// TIA Portal project "Hydroelectric Power Plant" (V20) (continued)
VERSION : 0.1
   VAR
      Os1 : Bool;
      Os2 : Bool;
      Os3 : Bool;
      Os4 : Bool;
      Os5 : Bool;
      Os6 : Bool;
      Os7 : Bool;
      Os8 : Bool;
      Os9 : Bool;
      Os10 : Bool;
      Os11 : Bool;
      Os12 : Bool;
   END_VAR
   VAR_TEMP   // added for the SCL form of the ladder/FBD networks
      _w1 : Bool;
      _w2 : Bool;
      _w3 : Bool;
   END_VAR
BEGIN

REGION Network 1
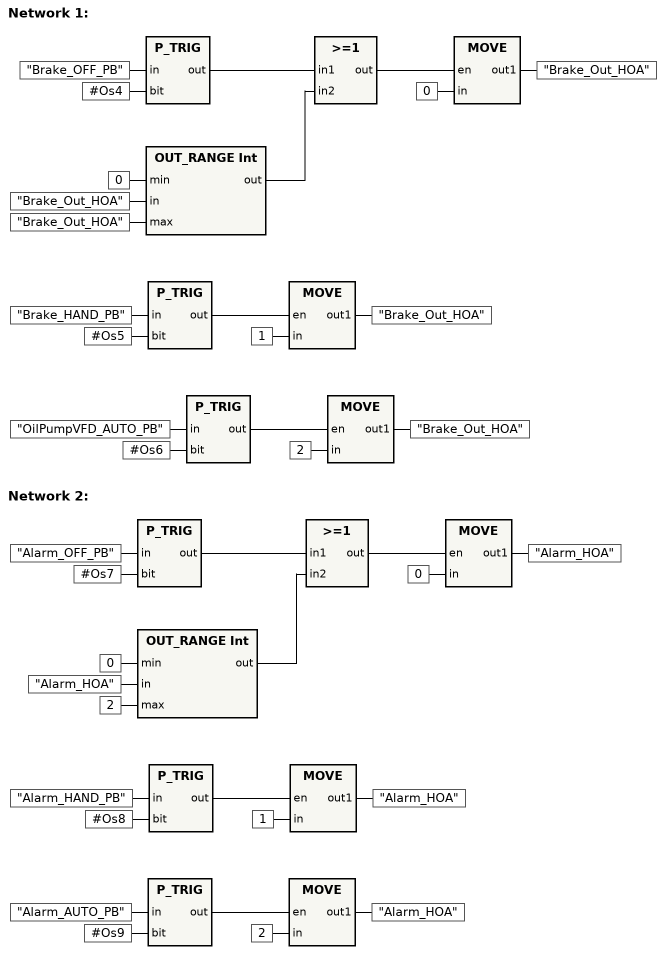
   #_w1 := "Brake_OFF_PB" AND NOT #Os4;   // rising edge
   #Os4 := "Brake_OFF_PB";
   IF #_w1 OR ("Brake_Out_HOA" < 0) OR ("Brake_Out_HOA" > "Brake_Out_HOA") THEN "Brake_Out_HOA" := 0; END_IF;
   #_w2 := "Brake_HAND_PB" AND NOT #Os5;   // rising edge
   #Os5 := "Brake_HAND_PB";
   IF #_w2 THEN "Brake_Out_HOA" := 1; END_IF;
   #_w3 := "OilPumpVFD_AUTO_PB" AND NOT #Os6;   // rising edge
   #Os6 := "OilPumpVFD_AUTO_PB";
   IF #_w3 THEN "Brake_Out_HOA" := 2; END_IF;
END_REGION

REGION Network 2
   #_w1 := "Alarm_OFF_PB" AND NOT #Os7;   // rising edge
   #Os7 := "Alarm_OFF_PB";
   IF #_w1 OR ("Alarm_HOA" < 0) OR ("Alarm_HOA" > 2) THEN "Alarm_HOA" := 0; END_IF;
   #_w2 := "Alarm_HAND_PB" AND NOT #Os8;   // rising edge
   #Os8 := "Alarm_HAND_PB";
   IF #_w2 THEN "Alarm_HOA" := 1; END_IF;
   #_w3 := "Alarm_AUTO_PB" AND NOT #Os9;   // rising edge
   #Os9 := "Alarm_AUTO_PB";
   IF #_w3 THEN "Alarm_HOA" := 2; END_IF;
END_REGION

REGION Network 3
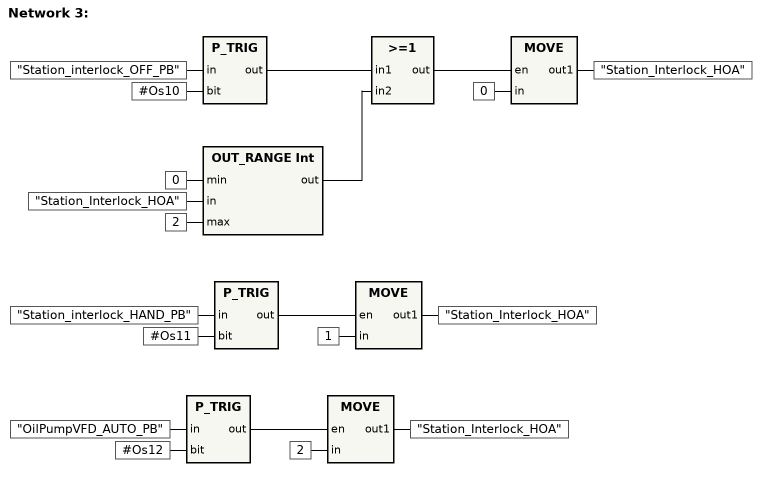
   #_w1 := "Station_interlock_OFF_PB" AND NOT #Os10;   // rising edge
   #Os10 := "Station_interlock_OFF_PB";
   IF #_w1 OR ("Station_Interlock_HOA" < 0) OR ("Station_Interlock_HOA" > 2) THEN
       "Station_Interlock_HOA" := 0;
   END_IF;
   #_w2 := "Station_interlock_HAND_PB" AND NOT #Os11;   // rising edge
   #Os11 := "Station_interlock_HAND_PB";
   IF #_w2 THEN "Station_Interlock_HOA" := 1; END_IF;
   #_w3 := "OilPumpVFD_AUTO_PB" AND NOT #Os12;   // rising edge
   #Os12 := "OilPumpVFD_AUTO_PB";
   IF #_w3 THEN "Station_Interlock_HOA" := 2; END_IF;
END_REGION
END_FUNCTION_BLOCK

FUNCTION_BLOCK "Alarm_FBD"   // FB11, FBD
{ S7_Optimized_Access := 'TRUE' }
VERSION : 0.1
   VAR
      OS1 : Bool;
      OS2 : Bool;
      OS3 : Bool;
      OS4 : Bool;
      OS5 : Bool;
      OS6 : Bool;
      OS7 : Bool;
      on8 : Bool;
   END_VAR
   VAR_TEMP
      tp1 : Int;
      OLFD : Time;
      tp2 : Int;
      OCD : Time;
      tp3 : Int;
      tp4 : Int;
      tp5 : Int;
      tp6 : Int;
      tp7 : Int;
      HOT : Time;
      OHF : Time;
      ROS : Time;
      BF : Time;
      AlarmTrigger : Bool;
   END_VAR
   VAR_TEMP   // added for the SCL form of the ladder/FBD networks
      _w1 : Bool;
   END_VAR
BEGIN

REGION Network 1: Oil_Low_Flow_Alarm
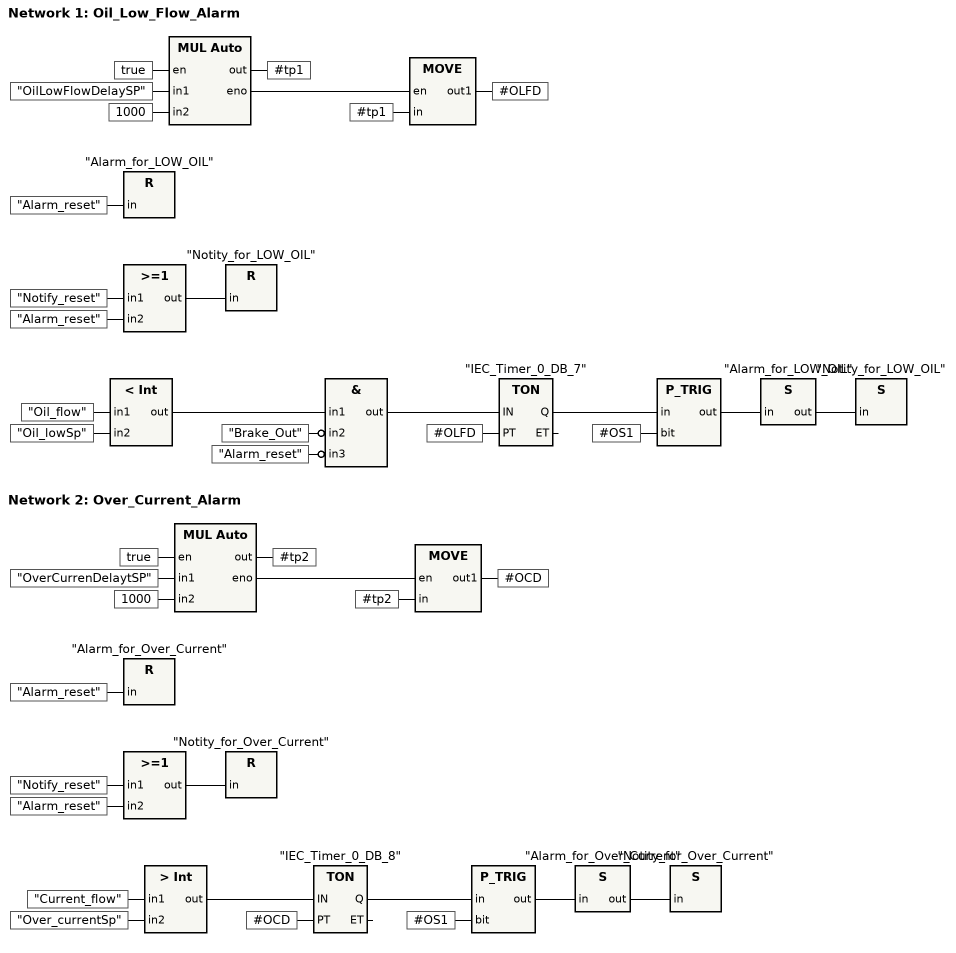
   IF true THEN
       #tp1 := "OilLowFlowDelaySP" * 1000;
       #OLFD := #tp1;
   END_IF;
   IF "Alarm_reset" THEN "Alarm_for_LOW_OIL" := FALSE; END_IF;
   IF "Notify_reset" OR "Alarm_reset" THEN "Notity_for_LOW_OIL" := FALSE; END_IF;
   "IEC_Timer_0_DB_7".TON(IN := ("Oil_flow" < "Oil_lowSp") AND NOT "Brake_Out" AND NOT "Alarm_reset",
                          PT := #OLFD);
   #_w1 := "IEC_Timer_0_DB_7".Q AND NOT #OS1;   // rising edge
   #OS1 := "IEC_Timer_0_DB_7".Q;
   IF #_w1 THEN
       "Alarm_for_LOW_OIL" := TRUE;
       "Notity_for_LOW_OIL" := TRUE;
   END_IF;
END_REGION

REGION Network 2: Over_Current_Alarm
   IF true THEN
       #tp2 := "OverCurrenDelaytSP" * 1000;
       #OCD := #tp2;
   END_IF;
   IF "Alarm_reset" THEN "Alarm_for_Over_Current" := FALSE; END_IF;
   IF "Notify_reset" OR "Alarm_reset" THEN "Notity_for_Over_Current" := FALSE; END_IF;
   "IEC_Timer_0_DB_8".TON(IN := "Current_flow" > "Over_currentSp", PT := #OCD);
   #_w1 := "IEC_Timer_0_DB_8".Q AND NOT #OS1;   // rising edge
   #OS1 := "IEC_Timer_0_DB_8".Q;
   IF #_w1 THEN
       "Alarm_for_Over_Current" := TRUE;
       "Notity_for_Over_Current" := TRUE;
   END_IF;
END_REGION

REGION Network 3: High_Oil_Temp_Alarm
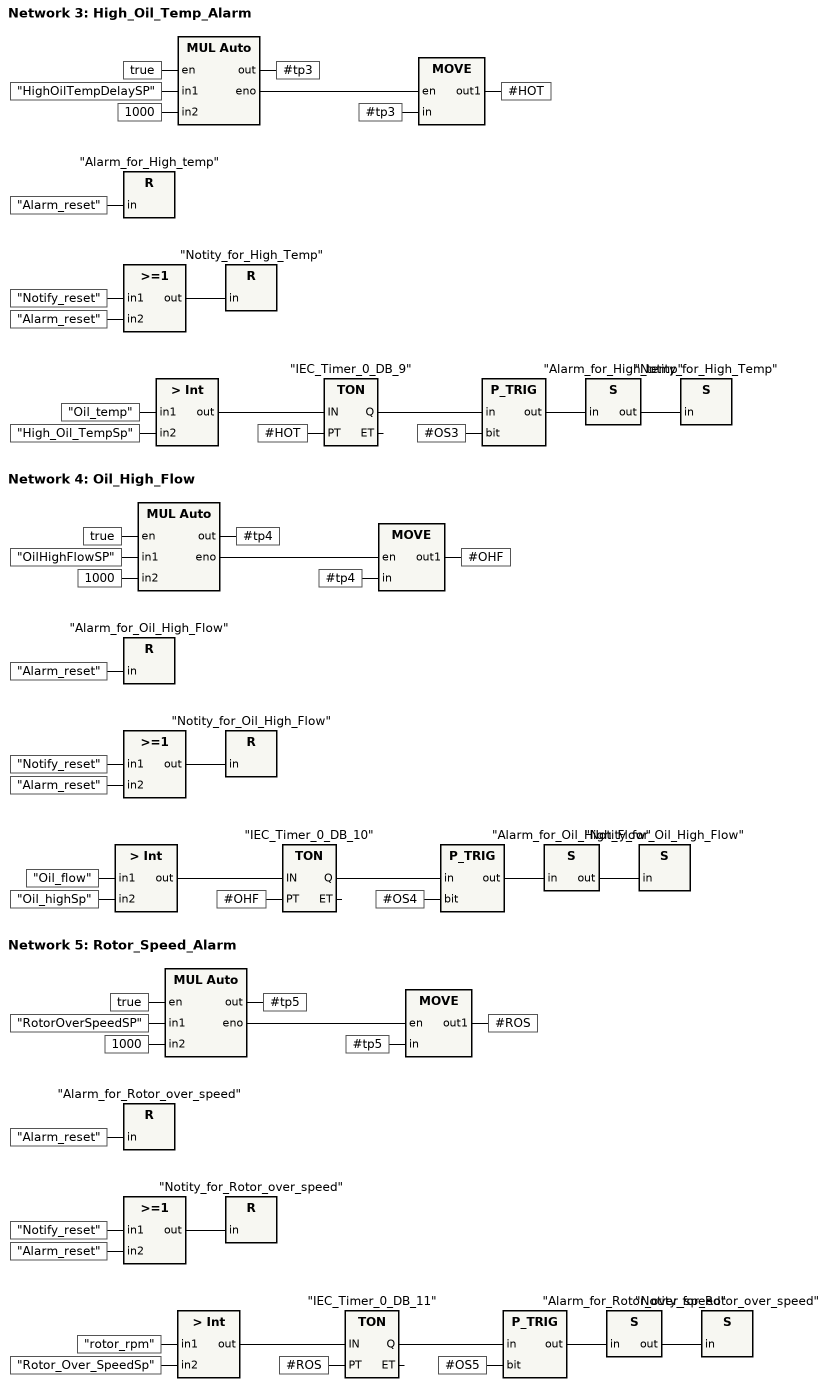
   IF true THEN
       #tp3 := "HighOilTempDelaySP" * 1000;
       #HOT := #tp3;
   END_IF;
   IF "Alarm_reset" THEN "Alarm_for_High_temp" := FALSE; END_IF;
   IF "Notify_reset" OR "Alarm_reset" THEN "Notity_for_High_Temp" := FALSE; END_IF;
   "IEC_Timer_0_DB_9".TON(IN := "Oil_temp" > "High_Oil_TempSp", PT := #HOT);
   #_w1 := "IEC_Timer_0_DB_9".Q AND NOT #OS3;   // rising edge
   #OS3 := "IEC_Timer_0_DB_9".Q;
   IF #_w1 THEN
       "Alarm_for_High_temp" := TRUE;
       "Notity_for_High_Temp" := TRUE;
   END_IF;
END_REGION

REGION Network 4: Oil_High_Flow
   IF true THEN
       #tp4 := "OilHighFlowSP" * 1000;
       #OHF := #tp4;
   END_IF;
   IF "Alarm_reset" THEN "Alarm_for_Oil_High_Flow" := FALSE; END_IF;
   IF "Notify_reset" OR "Alarm_reset" THEN "Notity_for_Oil_High_Flow" := FALSE; END_IF;
   "IEC_Timer_0_DB_10".TON(IN := "Oil_flow" > "Oil_highSp", PT := #OHF);
   #_w1 := "IEC_Timer_0_DB_10".Q AND NOT #OS4;   // rising edge
   #OS4 := "IEC_Timer_0_DB_10".Q;
   IF #_w1 THEN
       "Alarm_for_Oil_High_Flow" := TRUE;
       "Notity_for_Oil_High_Flow" := TRUE;
   END_IF;
END_REGION

REGION Network 5: Rotor_Speed_Alarm
   IF true THEN
       #tp5 := "RotorOverSpeedSP" * 1000;
       #ROS := #tp5;
   END_IF;
   IF "Alarm_reset" THEN "Alarm_for_Rotor_over_speed" := FALSE; END_IF;
   IF "Notify_reset" OR "Alarm_reset" THEN "Notity_for_Rotor_over_speed" := FALSE; END_IF;
   "IEC_Timer_0_DB_11".TON(IN := "rotor_rpm" > "Rotor_Over_SpeedSp", PT := #ROS);
   #_w1 := "IEC_Timer_0_DB_11".Q AND NOT #OS5;   // rising edge
   #OS5 := "IEC_Timer_0_DB_11".Q;
   IF #_w1 THEN
       "Alarm_for_Rotor_over_speed" := TRUE;
       "Notity_for_Rotor_over_speed" := TRUE;
   END_IF;
END_REGION

REGION Network 6: Brake_Failure_Alarm
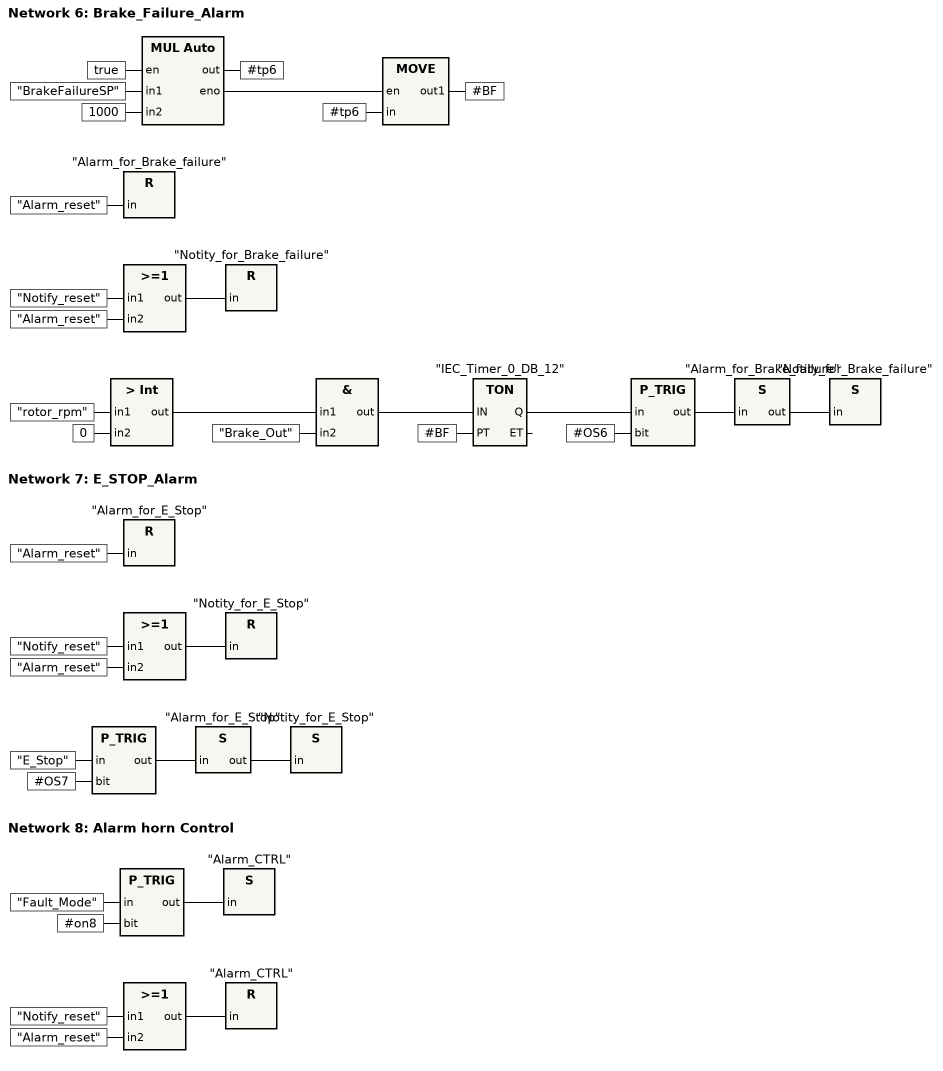
   IF true THEN
       #tp6 := "BrakeFailureSP" * 1000;
       #BF := #tp6;
   END_IF;
   IF "Alarm_reset" THEN "Alarm_for_Brake_failure" := FALSE; END_IF;
   IF "Notify_reset" OR "Alarm_reset" THEN "Notity_for_Brake_failure" := FALSE; END_IF;
   "IEC_Timer_0_DB_12".TON(IN := ("rotor_rpm" > 0) AND "Brake_Out", PT := #BF);
   #_w1 := "IEC_Timer_0_DB_12".Q AND NOT #OS6;   // rising edge
   #OS6 := "IEC_Timer_0_DB_12".Q;
   IF #_w1 THEN
       "Alarm_for_Brake_failure" := TRUE;
       "Notity_for_Brake_failure" := TRUE;
   END_IF;
END_REGION

REGION Network 7: E_STOP_Alarm
   IF "Alarm_reset" THEN "Alarm_for_E_Stop" := FALSE; END_IF;
   IF "Notify_reset" OR "Alarm_reset" THEN "Notity_for_E_Stop" := FALSE; END_IF;
   #_w1 := "E_Stop" AND NOT #OS7;   // rising edge
   #OS7 := "E_Stop";
   IF #_w1 THEN
       "Alarm_for_E_Stop" := TRUE;
       "Notity_for_E_Stop" := TRUE;
   END_IF;
END_REGION

REGION Network 8: Alarm horn Control
   #_w1 := "Fault_Mode" AND NOT #on8;   // rising edge
   #on8 := "Fault_Mode";
   IF #_w1 THEN "Alarm_CTRL" := TRUE; END_IF;
   IF "Notify_reset" OR "Alarm_reset" THEN "Alarm_CTRL" := FALSE; END_IF;
END_REGION
END_FUNCTION_BLOCK

FUNCTION_BLOCK "Modes_FBD"   // FB15, FBD
{ S7_Optimized_Access := 'TRUE' }
VERSION : 0.1
   VAR
      os1 : Bool;
      os2 : Bool;
      os3 : Bool;
      os4 : Bool;
      os5 : Bool;
      os6 : Bool;
   END_VAR
   VAR_TEMP
      ti1 : Time;
      tv2 : Int;
      tv1 : Int;
      ti2 : Time;
      ti3 : Time;
   END_VAR
   VAR_TEMP   // added for the SCL form of the ladder/FBD networks
      _w1 : Bool;
      _w2 : Bool;
      _w3 : Bool;
   END_VAR
BEGIN

REGION Network 1: WarmUp_Mode
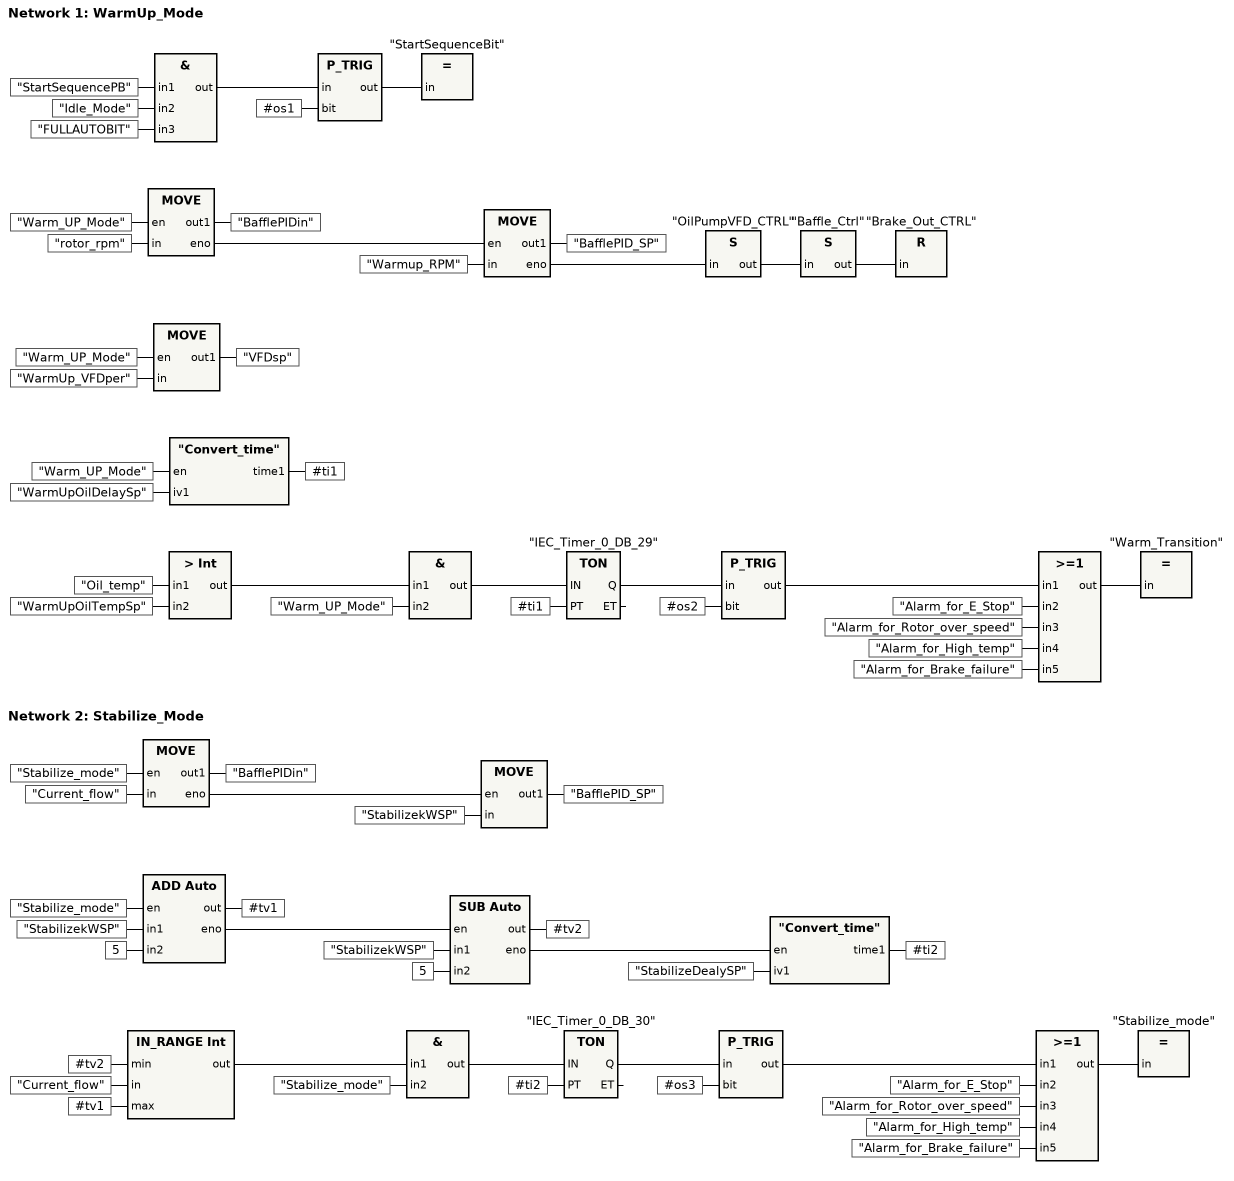
   #_w1 := "StartSequencePB" AND "Idle_Mode" AND "FULLAUTOBIT";
   #_w2 := #_w1 AND NOT #os1;   // rising edge
   #os1 := #_w1;
   "StartSequenceBit" := #_w2;
   IF "Warm_UP_Mode" THEN
       "BafflePIDin" := "rotor_rpm";
       "BafflePID_SP" := "Warmup_RPM";
       "OilPumpVFD_CTRL" := TRUE;
       "Baffle_Ctrl" := TRUE;
       "Brake_Out_CTRL" := FALSE;
       "VFDsp" := "WarmUp_VFDper";
       "Convert_time"(iv1 := "WarmUpOilDelaySp", time1 => #ti1);
   END_IF;
   "IEC_Timer_0_DB_29".TON(IN := ("Oil_temp" > "WarmUpOilTempSp") AND "Warm_UP_Mode", PT := #ti1);
   #_w3 := "IEC_Timer_0_DB_29".Q AND NOT #os2;   // rising edge
   #os2 := "IEC_Timer_0_DB_29".Q;
   "Warm_Transition" := #_w3 OR "Alarm_for_E_Stop" OR "Alarm_for_Rotor_over_speed" OR "Alarm_for_High_temp" OR "Alarm_for_Brake_failure";
END_REGION

REGION Network 2: Stabilize_Mode
   IF "Stabilize_mode" THEN
       "BafflePIDin" := "Current_flow";
       "BafflePID_SP" := "StabilizekWSP";
       #tv1 := "StabilizekWSP" + 5;
       #tv2 := "StabilizekWSP" - 5;
       "Convert_time"(iv1 := "StabilizeDealySP", time1 => #ti2);
   END_IF;
   "IEC_Timer_0_DB_30".TON(IN := (#tv2 <= "Current_flow") AND ("Current_flow" <= #tv1) AND "Stabilize_mode",
                           PT := #ti2);
   #_w1 := "IEC_Timer_0_DB_30".Q AND NOT #os3;   // rising edge
   #os3 := "IEC_Timer_0_DB_30".Q;
   "Stabilize_mode" := #_w1 OR "Alarm_for_E_Stop" OR "Alarm_for_Rotor_over_speed" OR "Alarm_for_High_temp" OR "Alarm_for_Brake_failure";
END_REGION

REGION Network 3: Gereration_Mode
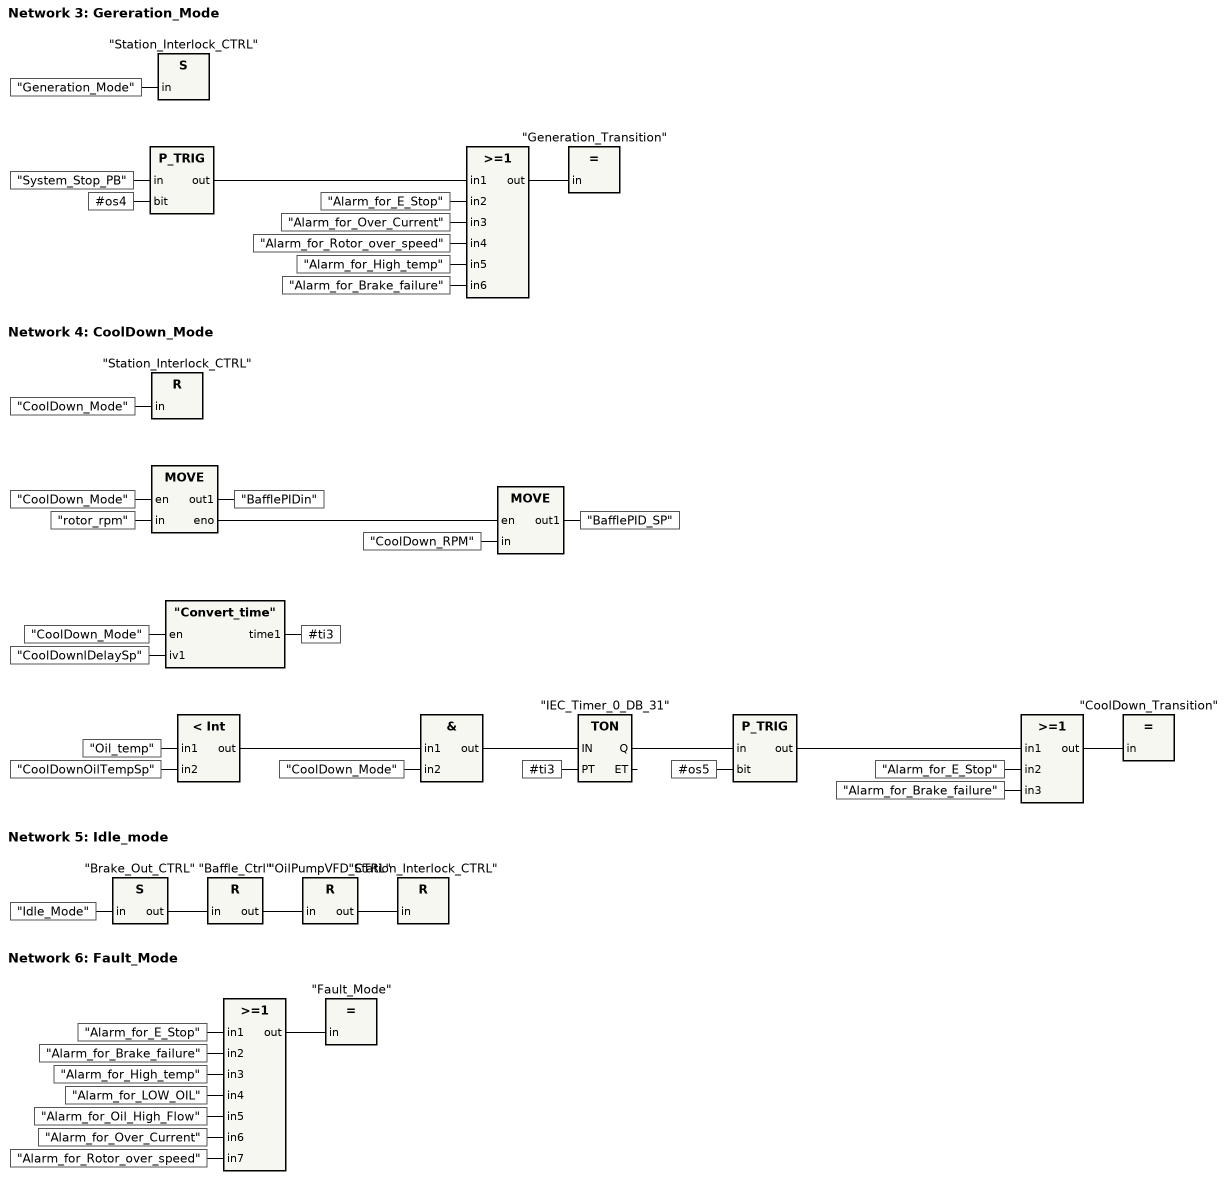
   IF "Generation_Mode" THEN "Station_Interlock_CTRL" := TRUE; END_IF;
   #_w1 := "System_Stop_PB" AND NOT #os4;   // rising edge
   #os4 := "System_Stop_PB";
   "Generation_Transition" := #_w1 OR "Alarm_for_E_Stop" OR "Alarm_for_Over_Current" OR "Alarm_for_Rotor_over_speed" OR "Alarm_for_High_temp" OR "Alarm_for_Brake_failure";
END_REGION

REGION Network 4: CoolDown_Mode
   IF "CoolDown_Mode" THEN
       "Station_Interlock_CTRL" := FALSE;
       "BafflePIDin" := "rotor_rpm";
       "BafflePID_SP" := "CoolDown_RPM";
       "Convert_time"(iv1 := "CoolDownlDelaySp", time1 => #ti3);
   END_IF;
   "IEC_Timer_0_DB_31".TON(IN := ("Oil_temp" < "CoolDownOilTempSp") AND "CoolDown_Mode", PT := #ti3);
   #_w1 := "IEC_Timer_0_DB_31".Q AND NOT #os5;   // rising edge
   #os5 := "IEC_Timer_0_DB_31".Q;
   "CoolDown_Transition" := #_w1 OR "Alarm_for_E_Stop" OR "Alarm_for_Brake_failure";
END_REGION

REGION Network 5: Idle_mode
   IF "Idle_Mode" THEN
       "Brake_Out_CTRL" := TRUE;
       "Baffle_Ctrl" := FALSE;
       "OilPumpVFD_CTRL" := FALSE;
       "Station_Interlock_CTRL" := FALSE;
   END_IF;
END_REGION

REGION Network 6: Fault_Mode
   "Fault_Mode" := "Alarm_for_E_Stop" OR "Alarm_for_Brake_failure" OR "Alarm_for_High_temp" OR "Alarm_for_LOW_OIL" OR "Alarm_for_Oil_High_Flow" OR "Alarm_for_Over_Current" OR "Alarm_for_Rotor_over_speed";
END_REGION
END_FUNCTION_BLOCK

FUNCTION_BLOCK "HOURMETER_FBD"   // FB20, FBD
{ S7_Optimized_Access := 'TRUE' }
VERSION : 0.1
   VAR
      Min_time_down : Bool;
      Min_countdown : Bool;
      Hour_countdown : Bool;
      Day_countdown : Bool;
      Day_count_down : Bool;
      Hr_count_down : Bool;
      reset_rto : Bool;
      min_count_reset : Bool;
      hour_count_reset : Bool;
      reset_hourmeter_trigger : Bool;
      os3 : Bool;
      os2 : Bool;
      os1 : Bool;
      os4 : Bool;
      Reset_HM_Trigger : Bool;
      accum_elapsed : Time;
   END_VAR
   VAR_TEMP
      resettime : Time;
   END_VAR
   VAR_TEMP   // added for the SCL form of the ladder/FBD networks
      _w1 : Bool;
      _w2 : Bool;
      _w3 : Bool;
   END_VAR
BEGIN

REGION Network 1
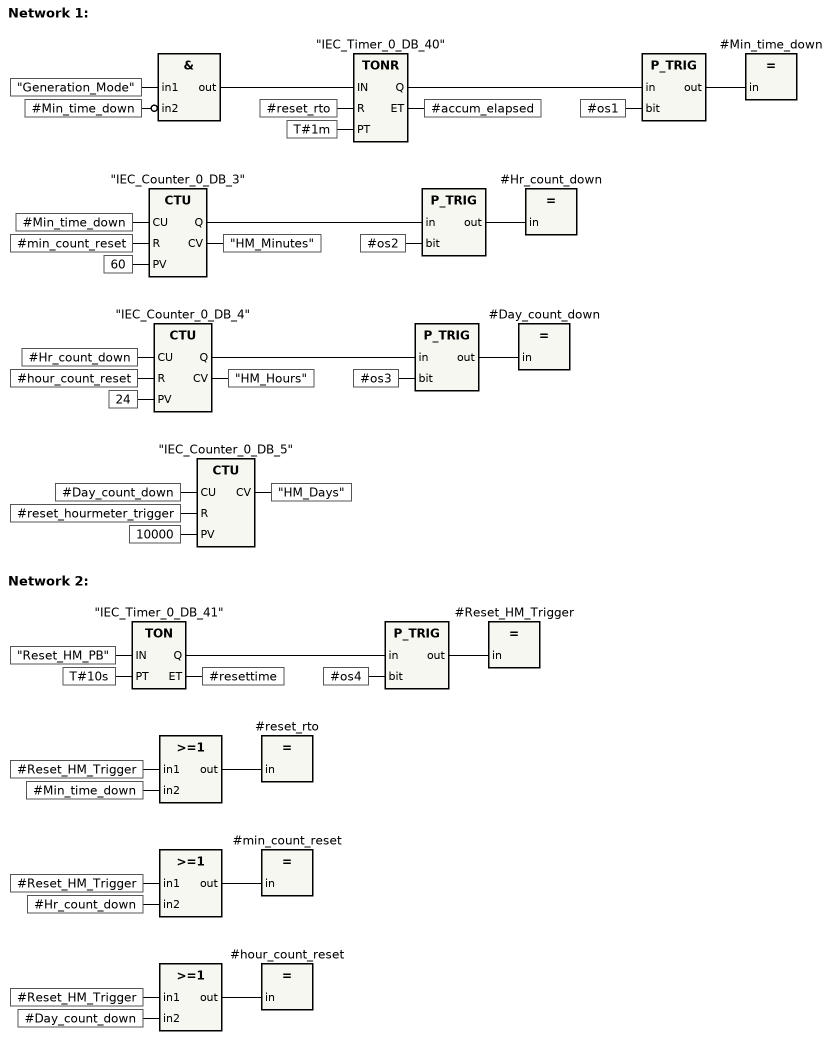
   "IEC_Timer_0_DB_40".TONR(IN := "Generation_Mode" AND NOT #Min_time_down,
                           R := #reset_rto,
                           PT := T#1m,
                           ET => #accum_elapsed);
   #_w1 := "IEC_Timer_0_DB_40".Q AND NOT #os1;   // rising edge
   #os1 := "IEC_Timer_0_DB_40".Q;
   #Min_time_down := #_w1;
   "IEC_Counter_0_DB_3".CTU(CU := #Min_time_down, R := #min_count_reset, PV := 60, CV => "HM_Minutes");
   #_w2 := "IEC_Counter_0_DB_3".Q AND NOT #os2;   // rising edge
   #os2 := "IEC_Counter_0_DB_3".Q;
   #Hr_count_down := #_w2;
   "IEC_Counter_0_DB_4".CTU(CU := #Hr_count_down, R := #hour_count_reset, PV := 24, CV => "HM_Hours");
   #_w3 := "IEC_Counter_0_DB_4".Q AND NOT #os3;   // rising edge
   #os3 := "IEC_Counter_0_DB_4".Q;
   #Day_count_down := #_w3;
   "IEC_Counter_0_DB_5".CTU(CU := #Day_count_down, R := #reset_hourmeter_trigger, PV := 10000, CV => "HM_Days");
END_REGION

REGION Network 2
   "IEC_Timer_0_DB_41".TON(IN := "Reset_HM_PB", PT := T#10s, ET => #resettime);
   #_w1 := "IEC_Timer_0_DB_41".Q AND NOT #os4;   // rising edge
   #os4 := "IEC_Timer_0_DB_41".Q;
   #Reset_HM_Trigger := #_w1;
   #reset_rto := #Reset_HM_Trigger OR #Min_time_down;
   #min_count_reset := #Reset_HM_Trigger OR #Hr_count_down;
   #hour_count_reset := #Reset_HM_Trigger OR #Day_count_down;
END_REGION
END_FUNCTION_BLOCK

// folder: LAD

FUNCTION_BLOCK "I/O LAD"   // FB2, LAD
{ S7_Optimized_Access := 'TRUE' }
VERSION : 0.1
// Gonna defined Analog and Digital I/O :p
BEGIN

REGION Network 1: Digital Output's
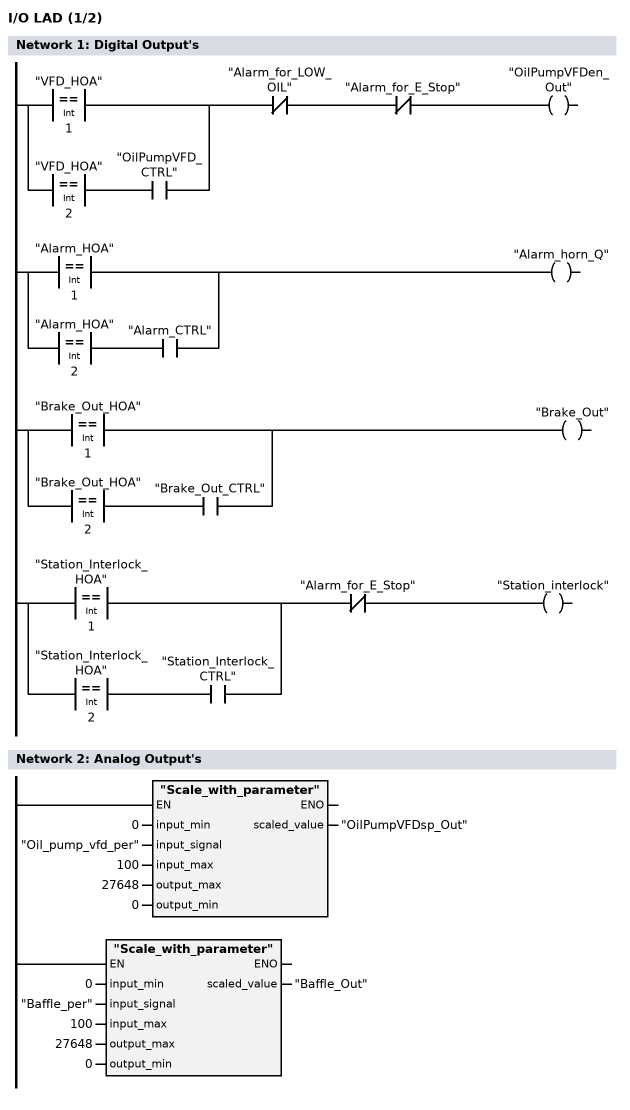
   RUNG wire#powerrail
      { S7_Templates := "SrcType := Int" } EQ_Contact(in1 := "VFD_HOA", in2 := 1)
      wire#w1
      I_Contact( "Alarm_for_LOW_OIL" )
      I_Contact( "Alarm_for_E_Stop" )
      Coil( "OilPumpVFDen_Out" )
   END_RUNG
   RUNG wire#powerrail
      { S7_Templates := "SrcType := Int" } EQ_Contact(in1 := "VFD_HOA", in2 := 2)
      Contact( "OilPumpVFD_CTRL" )
   END_RUNG wire#w1
   RUNG wire#powerrail
      { S7_Templates := "SrcType := Int" } EQ_Contact(in1 := "Alarm_HOA", in2 := 1)
      wire#w2
      Coil( "Alarm_horn_Q" )
   END_RUNG
   RUNG wire#powerrail
      { S7_Templates := "SrcType := Int" } EQ_Contact(in1 := "Alarm_HOA", in2 := 2)
      Contact( "Alarm_CTRL" )
   END_RUNG wire#w2
   RUNG wire#powerrail
      { S7_Templates := "SrcType := Int" } EQ_Contact(in1 := "Brake_Out_HOA", in2 := 1)
      wire#w3
      Coil( "Brake_Out" )
   END_RUNG
   RUNG wire#powerrail
      { S7_Templates := "SrcType := Int" } EQ_Contact(in1 := "Brake_Out_HOA", in2 := 2)
      Contact( "Brake_Out_CTRL" )
   END_RUNG wire#w3
   RUNG wire#powerrail
      { S7_Templates := "SrcType := Int" } EQ_Contact(in1 := "Station_Interlock_HOA", in2 := 1)
      wire#w4
      I_Contact( "Alarm_for_E_Stop" )
      Coil( "Station_interlock" )
   END_RUNG
   RUNG wire#powerrail
      { S7_Templates := "SrcType := Int" } EQ_Contact(in1 := "Station_Interlock_HOA", in2 := 2)
      Contact( "Station_Interlock_CTRL" )
   END_RUNG wire#w4
   // the same network as SCL:
   "OilPumpVFDen_Out" := (("VFD_HOA" = 1) OR (("VFD_HOA" = 2) AND "OilPumpVFD_CTRL")) AND NOT "Alarm_for_LOW_OIL" AND NOT "Alarm_for_E_Stop";
   "Alarm_horn_Q" := ("Alarm_HOA" = 1) OR (("Alarm_HOA" = 2) AND "Alarm_CTRL");
   "Brake_Out" := ("Brake_Out_HOA" = 1) OR (("Brake_Out_HOA" = 2) AND "Brake_Out_CTRL");
   "Station_interlock" := (("Station_Interlock_HOA" = 1) OR (("Station_Interlock_HOA" = 2) AND "Station_Interlock_CTRL")) AND NOT "Alarm_for_E_Stop";
END_REGION

REGION Network 2: Analog Output's
   RUNG wire#powerrail
      "Scale_with_parameter"(input_min := 0, input_signal := "Oil_pump_vfd_per", input_max := 100, output_max := 27648, output_min := 0, scaled_value => "OilPumpVFDsp_Out")
   END_RUNG
   RUNG wire#powerrail
      "Scale_with_parameter"(input_min := 0, input_signal := "Baffle_per", input_max := 100, output_max := 27648, output_min := 0, scaled_value => "Baffle_Out")
   END_RUNG
   // the same network as SCL:
   "Scale_with_parameter"(input_min := 0,
                          input_signal := "Oil_pump_vfd_per",
                          input_max := 100,
                          output_max := 27648,
                          output_min := 0,
                          scaled_value => "OilPumpVFDsp_Out");
   "Scale_with_parameter"(input_min := 0,
                          input_signal := "Baffle_per",
                          input_max := 100,
                          output_max := 27648,
                          output_min := 0,
                          scaled_value => "Baffle_Out");
END_REGION

REGION Network 3: Analog Input's
